   hmiStns[1].wip[14].pnCode[4] := 0;
   hmiStns[1].wip[14].pnCode[5] := 0;
   hmiStns[1].wip[14].pnCode[6] := 0;
   hmiStns[1].wip[14].pnCode[7] := 0;
   hmiStns[1].wip[15].wipCode := -1;
   hmiStns[1].wip[15].pnCode[0] := 0;
   hmiStns[1].wip[15].pnCode[1] := 0;
   hmiStns[1].wip[15].pnCode[2] := 0;
   hmiStns[1].wip[15].pnCode[3] := 0;
   hmiStns[1].wip[15].pnCode[4] := 0;
   hmiStns[1].wip[15].pnCode[5] := 0;
   hmiStns[1].wip[15].pnCode[6] := 0;
   hmiStns[1].wip[15].pnCode[7] := 0;
   hmiStns[1].wip[16].wipCode := -1;
   hmiStns[1].wip[16].pnCode[0] := 0;
   hmiStns[1].wip[16].pnCode[1] := 0;
   hmiStns[1].wip[16].pnCode[2] := 0;
   hmiStns[1].wip[16].pnCode[3] := 0;
   hmiStns[1].wip[16].pnCode[4] := 0;
   hmiStns[1].wip[16].pnCode[5] := 0;
   hmiStns[1].wip[16].pnCode[6] := 0;
   hmiStns[1].wip[16].pnCode[7] := 0;
   hmiStns[1].wip[17].wipCode := -1;
   hmiStns[1].wip[17].pnCode[0] := 0;
   hmiStns[1].wip[17].pnCode[1] := 0;
   hmiStns[1].wip[17].pnCode[2] := 0;
   hmiStns[1].wip[17].pnCode[3] := 0;
   hmiStns[1].wip[17].pnCode[4] := 0;
   hmiStns[1].wip[17].pnCode[5] := 0;
   hmiStns[1].wip[17].pnCode[6] := 0;
   hmiStns[1].wip[17].pnCode[7] := 0;
   hmiStns[1].wip[18].wipCode := -1;
   hmiStns[1].wip[18].pnCode[0] := 0;
   hmiStns[1].wip[18].pnCode[1] := 0;
   hmiStns[1].wip[18].pnCode[2] := 0;
   hmiStns[1].wip[18].pnCode[3] := 0;
   hmiStns[1].wip[18].pnCode[4] := 0;
   hmiStns[1].wip[18].pnCode[5] := 0;
   hmiStns[1].wip[18].pnCode[6] := 0;
   hmiStns[1].wip[18].pnCode[7] := 0;
   hmiStns[1].wip[19].wipCode := -1;
   hmiStns[1].wip[19].pnCode[0] := 0;
   hmiStns[1].wip[19].pnCode[1] := 0;
   hmiStns[1].wip[19].pnCode[2] := 0;
   hmiStns[1].wip[19].pnCode[3] := 0;
   hmiStns[1].wip[19].pnCode[4] := 0;
   hmiStns[1].wip[19].pnCode[5] := 0;
   hmiStns[1].wip[19].pnCode[6] := 0;
   hmiStns[1].wip[19].pnCode[7] := 0;
   hmiStns[1].wip[20].wipCode := -1;
   hmiStns[1].wip[20].pnCode[0] := 0;
   hmiStns[1].wip[20].pnCode[1] := 0;
   hmiStns[1].wip[20].pnCode[2] := 0;
   hmiStns[1].wip[20].pnCode[3] := 0;
   hmiStns[1].wip[20].pnCode[4] := 0;
   hmiStns[1].wip[20].pnCode[5] := 0;
   hmiStns[1].wip[20].pnCode[6] := 0;
   hmiStns[1].wip[20].pnCode[7] := 0;
   hmiStns[1].wip[21].wipCode := -1;
   hmiStns[1].wip[21].pnCode[0] := 0;
   hmiStns[1].wip[21].pnCode[1] := 0;
   hmiStns[1].wip[21].pnCode[2] := 0;
   hmiStns[1].wip[21].pnCode[3] := 0;
   hmiStns[1].wip[21].pnCode[4] := 0;
   hmiStns[1].wip[21].pnCode[5] := 0;
   hmiStns[1].wip[21].pnCode[6] := 0;
   hmiStns[1].wip[21].pnCode[7] := 0;
   hmiStns[1].wip[22].wipCode := -1;
   hmiStns[1].wip[22].pnCode[0] := 0;
   hmiStns[1].wip[22].pnCode[1] := 0;
   hmiStns[1].wip[22].pnCode[2] := 0;
   hmiStns[1].wip[22].pnCode[3] := 0;
   hmiStns[1].wip[22].pnCode[4] := 0;
   hmiStns[1].wip[22].pnCode[5] := 0;
   hmiStns[1].wip[22].pnCode[6] := 0;
   hmiStns[1].wip[22].pnCode[7] := 0;
   hmiStns[1].wip[23].wipCode := -1;
   hmiStns[1].wip[23].pnCode[0] := 0;
   hmiStns[1].wip[23].pnCode[1] := 0;
   hmiStns[1].wip[23].pnCode[2] := 0;
   hmiStns[1].wip[23].pnCode[3] := 0;
   hmiStns[1].wip[23].pnCode[4] := 0;
   hmiStns[1].wip[23].pnCode[5] := 0;
   hmiStns[1].wip[23].pnCode[6] := 0;
   hmiStns[1].wip[23].pnCode[7] := 0;
   hmiStns[1].wip[24].wipCode := -1;
   hmiStns[1].wip[24].pnCode[0] := 0;
   hmiStns[1].wip[24].pnCode[1] := 0;
   hmiStns[1].wip[24].pnCode[2] := 0;
   hmiStns[1].wip[24].pnCode[3] := 0;
   hmiStns[1].wip[24].pnCode[4] := 0;
   hmiStns[1].wip[24].pnCode[5] := 0;
   hmiStns[1].wip[24].pnCode[6] := 0;
   hmiStns[1].wip[24].pnCode[7] := 0;
   hmiStns[1].wip[25].wipCode := -1;
   hmiStns[1].wip[25].pnCode[0] := 0;
   hmiStns[1].wip[25].pnCode[1] := 0;
   hmiStns[1].wip[25].pnCode[2] := 0;
   hmiStns[1].wip[25].pnCode[3] := 0;
   hmiStns[1].wip[25].pnCode[4] := 0;
   hmiStns[1].wip[25].pnCode[5] := 0;
   hmiStns[1].wip[25].pnCode[6] := 0;
   hmiStns[1].wip[25].pnCode[7] := 0;
   hmiStns[1].wip[26].wipCode := -1;
   hmiStns[1].wip[26].pnCode[0] := 0;
   hmiStns[1].wip[26].pnCode[1] := 0;
   hmiStns[1].wip[26].pnCode[2] := 0;
   hmiStns[1].wip[26].pnCode[3] := 0;
   hmiStns[1].wip[26].pnCode[4] := 0;
   hmiStns[1].wip[26].pnCode[5] := 0;
   hmiStns[1].wip[26].pnCode[6] := 0;
   hmiStns[1].wip[26].pnCode[7] := 0;
   hmiStns[1].wip[27].wipCode := -1;
   hmiStns[1].wip[27].pnCode[0] := 0;
   hmiStns[1].wip[27].pnCode[1] := 0;
   hmiStns[1].wip[27].pnCode[2] := 0;
   hmiStns[1].wip[27].pnCode[3] := 0;
   hmiStns[1].wip[27].pnCode[4] := 0;
   hmiStns[1].wip[27].pnCode[5] := 0;
   hmiStns[1].wip[27].pnCode[6] := 0;
   hmiStns[1].wip[27].pnCode[7] := 0;
   hmiStns[1].wip[28].wipCode := -1;
   hmiStns[1].wip[28].pnCode[0] := 0;
   hmiStns[1].wip[28].pnCode[1] := 0;
   hmiStns[1].wip[28].pnCode[2] := 0;
   hmiStns[1].wip[28].pnCode[3] := 0;
   hmiStns[1].wip[28].pnCode[4] := 0;
   hmiStns[1].wip[28].pnCode[5] := 0;
   hmiStns[1].wip[28].pnCode[6] := 0;
   hmiStns[1].wip[28].pnCode[7] := 0;
   hmiStns[1].wip[29].wipCode := -1;
   hmiStns[1].wip[29].pnCode[0] := 0;
   hmiStns[1].wip[29].pnCode[1] := 0;
   hmiStns[1].wip[29].pnCode[2] := 0;
   hmiStns[1].wip[29].pnCode[3] := 0;
   hmiStns[1].wip[29].pnCode[4] := 0;
   hmiStns[1].wip[29].pnCode[5] := 0;
   hmiStns[1].wip[29].pnCode[6] := 0;
   hmiStns[1].wip[29].pnCode[7] := 0;
   hmiStns[1].wip[30].wipCode := -1;
   hmiStns[1].wip[30].pnCode[0] := 0;
   hmiStns[1].wip[30].pnCode[1] := 0;
   hmiStns[1].wip[30].pnCode[2] := 0;
   hmiStns[1].wip[30].pnCode[3] := 0;
   hmiStns[1].wip[30].pnCode[4] := 0;
   hmiStns[1].wip[30].pnCode[5] := 0;
   hmiStns[1].wip[30].pnCode[6] := 0;
   hmiStns[1].wip[30].pnCode[7] := 0;
   hmiStns[1].wip[31].wipCode := -1;
   hmiStns[1].wip[31].pnCode[0] := 0;
   hmiStns[1].wip[31].pnCode[1] := 0;
   hmiStns[1].wip[31].pnCode[2] := 0;
   hmiStns[1].wip[31].pnCode[3] := 0;
   hmiStns[1].wip[31].pnCode[4] := 0;
   hmiStns[1].wip[31].pnCode[5] := 0;
   hmiStns[1].wip[31].pnCode[6] := 0;
   hmiStns[1].wip[31].pnCode[7] := 0;
   hmiStns[1].wip[32].wipCode := -1;
   hmiStns[1].wip[32].pnCode[0] := 0;
   hmiStns[1].wip[32].pnCode[1] := 0;
   hmiStns[1].wip[32].pnCode[2] := 0;
   hmiStns[1].wip[32].pnCode[3] := 0;
   hmiStns[1].wip[32].pnCode[4] := 0;
   hmiStns[1].wip[32].pnCode[5] := 0;
   hmiStns[1].wip[32].pnCode[6] := 0;
   hmiStns[1].wip[32].pnCode[7] := 0;
   hmiStns[1].wip[33].wipCode := -1;
   hmiStns[1].wip[33].pnCode[0] := 0;
   hmiStns[1].wip[33].pnCode[1] := 0;
   hmiStns[1].wip[33].pnCode[2] := 0;
   hmiStns[1].wip[33].pnCode[3] := 0;
   hmiStns[1].wip[33].pnCode[4] := 0;
   hmiStns[1].wip[33].pnCode[5] := 0;
   hmiStns[1].wip[33].pnCode[6] := 0;
   hmiStns[1].wip[33].pnCode[7] := 0;
   hmiStns[1].wip[34].wipCode := -1;
   hmiStns[1].wip[34].pnCode[0] := 0;
   hmiStns[1].wip[34].pnCode[1] := 0;
   hmiStns[1].wip[34].pnCode[2] := 0;
   hmiStns[1].wip[34].pnCode[3] := 0;
   hmiStns[1].wip[34].pnCode[4] := 0;
   hmiStns[1].wip[34].pnCode[5] := 0;
   hmiStns[1].wip[34].pnCode[6] := 0;
   hmiStns[1].wip[34].pnCode[7] := 0;
   hmiStns[1].wip[35].wipCode := -1;
   hmiStns[1].wip[35].pnCode[0] := 0;
   hmiStns[1].wip[35].pnCode[1] := 0;
   hmiStns[1].wip[35].pnCode[2] := 0;
   hmiStns[1].wip[35].pnCode[3] := 0;
   hmiStns[1].wip[35].pnCode[4] := 0;
   hmiStns[1].wip[35].pnCode[5] := 0;
   hmiStns[1].wip[35].pnCode[6] := 0;
   hmiStns[1].wip[35].pnCode[7] := 0;
   hmiStns[1].wip[36].wipCode := -1;
   hmiStns[1].wip[36].pnCode[0] := 0;
   hmiStns[1].wip[36].pnCode[1] := 0;
   hmiStns[1].wip[36].pnCode[2] := 0;
   hmiStns[1].wip[36].pnCode[3] := 0;
   hmiStns[1].wip[36].pnCode[4] := 0;
   hmiStns[1].wip[36].pnCode[5] := 0;
   hmiStns[1].wip[36].pnCode[6] := 0;
   hmiStns[1].wip[36].pnCode[7] := 0;
   hmiStns[1].wip[37].wipCode := -1;
   hmiStns[1].wip[37].pnCode[0] := 0;
   hmiStns[1].wip[37].pnCode[1] := 0;
   hmiStns[1].wip[37].pnCode[2] := 0;
   hmiStns[1].wip[37].pnCode[3] := 0;
   hmiStns[1].wip[37].pnCode[4] := 0;
   hmiStns[1].wip[37].pnCode[5] := 0;
   hmiStns[1].wip[37].pnCode[6] := 0;
   hmiStns[1].wip[37].pnCode[7] := 0;
   hmiStns[1].wip[38].wipCode := -1;
   hmiStns[1].wip[38].pnCode[0] := 0;
   hmiStns[1].wip[38].pnCode[1] := 0;
   hmiStns[1].wip[38].pnCode[2] := 0;
   hmiStns[1].wip[38].pnCode[3] := 0;
   hmiStns[1].wip[38].pnCode[4] := 0;
   hmiStns[1].wip[38].pnCode[5] := 0;
   hmiStns[1].wip[38].pnCode[6] := 0;
   hmiStns[1].wip[38].pnCode[7] := 0;
   hmiStns[1].wip[39].wipCode := -1;
   hmiStns[1].wip[39].pnCode[0] := 0;
   hmiStns[1].wip[39].pnCode[1] := 0;
   hmiStns[1].wip[39].pnCode[2] := 0;
   hmiStns[1].wip[39].pnCode[3] := 0;
   hmiStns[1].wip[39].pnCode[4] := 0;
   hmiStns[1].wip[39].pnCode[5] := 0;
   hmiStns[1].wip[39].pnCode[6] := 0;
   hmiStns[1].wip[39].pnCode[7] := 0;
   hmiStns[1].wip[40].wipCode := -1;
   hmiStns[1].wip[40].pnCode[0] := 0;
   hmiStns[1].wip[40].pnCode[1] := 0;
   hmiStns[1].wip[40].pnCode[2] := 0;
   hmiStns[1].wip[40].pnCode[3] := 0;
   hmiStns[1].wip[40].pnCode[4] := 0;
   hmiStns[1].wip[40].pnCode[5] := 0;
   hmiStns[1].wip[40].pnCode[6] := 0;
   hmiStns[1].wip[40].pnCode[7] := 0;
   hmiStns[1].wip[41].wipCode := -1;
   hmiStns[1].wip[41].pnCode[0] := 0;
   hmiStns[1].wip[41].pnCode[1] := 0;
   hmiStns[1].wip[41].pnCode[2] := 0;
   hmiStns[1].wip[41].pnCode[3] := 0;
   hmiStns[1].wip[41].pnCode[4] := 0;
   hmiStns[1].wip[41].pnCode[5] := 0;
   hmiStns[1].wip[41].pnCode[6] := 0;
   hmiStns[1].wip[41].pnCode[7] := 0;
   hmiStns[1].wip[42].wipCode := -1;
   hmiStns[1].wip[42].pnCode[0] := 0;
   hmiStns[1].wip[42].pnCode[1] := 0;
   hmiStns[1].wip[42].pnCode[2] := 0;
   hmiStns[1].wip[42].pnCode[3] := 0;
   hmiStns[1].wip[42].pnCode[4] := 0;
   hmiStns[1].wip[42].pnCode[5] := 0;
   hmiStns[1].wip[42].pnCode[6] := 0;
   hmiStns[1].wip[42].pnCode[7] := 0;
   hmiStns[1].wip[43].wipCode := -1;
   hmiStns[1].wip[43].pnCode[0] := 0;
   hmiStns[1].wip[43].pnCode[1] := 0;
   hmiStns[1].wip[43].pnCode[2] := 0;
   hmiStns[1].wip[43].pnCode[3] := 0;
   hmiStns[1].wip[43].pnCode[4] := 0;
   hmiStns[1].wip[43].pnCode[5] := 0;
   hmiStns[1].wip[43].pnCode[6] := 0;
   hmiStns[1].wip[43].pnCode[7] := 0;
   hmiStns[1].wip[44].wipCode := -1;
   hmiStns[1].wip[44].pnCode[0] := 0;
   hmiStns[1].wip[44].pnCode[1] := 0;
   hmiStns[1].wip[44].pnCode[2] := 0;
   hmiStns[1].wip[44].pnCode[3] := 0;
   hmiStns[1].wip[44].pnCode[4] := 0;
   hmiStns[1].wip[44].pnCode[5] := 0;
   hmiStns[1].wip[44].pnCode[6] := 0;
   hmiStns[1].wip[44].pnCode[7] := 0;
   hmiStns[1].wip[45].wipCode := -1;
   hmiStns[1].wip[45].pnCode[0] := 0;
   hmiStns[1].wip[45].pnCode[1] := 0;
   hmiStns[1].wip[45].pnCode[2] := 0;
   hmiStns[1].wip[45].pnCode[3] := 0;
   hmiStns[1].wip[45].pnCode[4] := 0;
   hmiStns[1].wip[45].pnCode[5] := 0;
   hmiStns[1].wip[45].pnCode[6] := 0;
   hmiStns[1].wip[45].pnCode[7] := 0;
   hmiStns[1].wip[46].wipCode := -1;
   hmiStns[1].wip[46].pnCode[0] := 0;
   hmiStns[1].wip[46].pnCode[1] := 0;
   hmiStns[1].wip[46].pnCode[2] := 0;
   hmiStns[1].wip[46].pnCode[3] := 0;
   hmiStns[1].wip[46].pnCode[4] := 0;
   hmiStns[1].wip[46].pnCode[5] := 0;
   hmiStns[1].wip[46].pnCode[6] := 0;
   hmiStns[1].wip[46].pnCode[7] := 0;
   hmiStns[1].wip[47].wipCode := -1;
   hmiStns[1].wip[47].pnCode[0] := 0;
   hmiStns[1].wip[47].pnCode[1] := 0;
   hmiStns[1].wip[47].pnCode[2] := 0;
   hmiStns[1].wip[47].pnCode[3] := 0;
   hmiStns[1].wip[47].pnCode[4] := 0;
   hmiStns[1].wip[47].pnCode[5] := 0;
   hmiStns[1].wip[47].pnCode[6] := 0;
   hmiStns[1].wip[47].pnCode[7] := 0;
   hmiStns[1].wip[48].wipCode := -1;
   hmiStns[1].wip[48].pnCode[0] := 0;
   hmiStns[1].wip[48].pnCode[1] := 0;
   hmiStns[1].wip[48].pnCode[2] := 0;
   hmiStns[1].wip[48].pnCode[3] := 0;
   hmiStns[1].wip[48].pnCode[4] := 0;
   hmiStns[1].wip[48].pnCode[5] := 0;
   hmiStns[1].wip[48].pnCode[6] := 0;
   hmiStns[1].wip[48].pnCode[7] := 0;
   hmiStns[1].wip[49].wipCode := -1;
   hmiStns[1].wip[49].pnCode[0] := 0;
   hmiStns[1].wip[49].pnCode[1] := 0;
   hmiStns[1].wip[49].pnCode[2] := 0;
   hmiStns[1].wip[49].pnCode[3] := 0;
   hmiStns[1].wip[49].pnCode[4] := 0;
   hmiStns[1].wip[49].pnCode[5] := 0;
   hmiStns[1].wip[49].pnCode[6] := 0;
   hmiStns[1].wip[49].pnCode[7] := 0;
   hmiStns[2].wip[0].wipCode := 53014;
   hmiStns[2].wip[0].pnCode[0] := 0;
   hmiStns[2].wip[0].pnCode[1] := 243000;
   hmiStns[2].wip[0].pnCode[2] := 148000;
   hmiStns[2].wip[0].pnCode[3] := 0;
   hmiStns[2].wip[0].pnCode[4] := 0;
   hmiStns[2].wip[0].pnCode[5] := 0;
   hmiStns[2].wip[0].pnCode[6] := 147000;
   hmiStns[2].wip[0].pnCode[7] := 149000;
   hmiStns[2].wip[1].wipCode := 19031;
   hmiStns[2].wip[1].pnCode[0] := 0;
   hmiStns[2].wip[1].pnCode[1] := 243000;
   hmiStns[2].wip[1].pnCode[2] := 53000;
   hmiStns[2].wip[1].pnCode[3] := 0;
   hmiStns[2].wip[1].pnCode[4] := 0;
   hmiStns[2].wip[1].pnCode[5] := 0;
   hmiStns[2].wip[1].pnCode[6] := 31000;
   hmiStns[2].wip[1].pnCode[7] := 71000;
   hmiStns[2].wip[2].wipCode := 21028;
   hmiStns[2].wip[2].pnCode[0] := 0;
   hmiStns[2].wip[2].pnCode[1] := 243000;
   hmiStns[2].wip[2].pnCode[2] := 57000;
   hmiStns[2].wip[2].pnCode[3] := 0;
   hmiStns[2].wip[2].pnCode[4] := 0;
   hmiStns[2].wip[2].pnCode[5] := 0;
   hmiStns[2].wip[2].pnCode[6] := 25000;
   hmiStns[2].wip[2].pnCode[7] := 18000;
   hmiStns[2].wip[3].wipCode := 22008;
   hmiStns[2].wip[3].pnCode[0] := 0;
   hmiStns[2].wip[3].pnCode[1] := 243000;
   hmiStns[2].wip[3].pnCode[2] := 84000;
   hmiStns[2].wip[3].pnCode[3] := 0;
   hmiStns[2].wip[3].pnCode[4] := 0;
   hmiStns[2].wip[3].pnCode[5] := 0;
   hmiStns[2].wip[3].pnCode[6] := 31000;
   hmiStns[2].wip[3].pnCode[7] := 71000;
   hmiStns[2].wip[4].wipCode := 20050;
   hmiStns[2].wip[4].pnCode[0] := 0;
   hmiStns[2].wip[4].pnCode[1] := 243000;
   hmiStns[2].wip[4].pnCode[2] := 70000;
   hmiStns[2].wip[4].pnCode[3] := 72000;
   hmiStns[2].wip[4].pnCode[4] := 0;
   hmiStns[2].wip[4].pnCode[5] := 58000;
   hmiStns[2].wip[4].pnCode[6] := 33000;
   hmiStns[2].wip[4].pnCode[7] := 73000;
   hmiStns[2].wip[5].wipCode := 27040;
   hmiStns[2].wip[5].pnCode[0] := 0;
   hmiStns[2].wip[5].pnCode[1] := 243000;
   hmiStns[2].wip[5].pnCode[2] := 127000;
   hmiStns[2].wip[5].pnCode[3] := 0;
   hmiStns[2].wip[5].pnCode[4] := 0;
   hmiStns[2].wip[5].pnCode[5] := 100000;
   hmiStns[2].wip[5].pnCode[6] := 101000;
   hmiStns[2].wip[5].pnCode[7] := 128000;
   hmiStns[2].wip[6].wipCode := 28041;
   hmiStns[2].wip[6].pnCode[0] := 0;
   hmiStns[2].wip[6].pnCode[1] := 243000;
   hmiStns[2].wip[6].pnCode[2] := 122000;
   hmiStns[2].wip[6].pnCode[3] := 123000;
   hmiStns[2].wip[6].pnCode[4] := 0;
   hmiStns[2].wip[6].pnCode[5] := 102000;
   hmiStns[2].wip[6].pnCode[6] := 103000;
   hmiStns[2].wip[6].pnCode[7] := 133000;
   hmiStns[2].wip[7].wipCode := 29044;
   hmiStns[2].wip[7].pnCode[0] := 0;
   hmiStns[2].wip[7].pnCode[1] := 243000;
   hmiStns[2].wip[7].pnCode[2] := 100000;
   hmiStns[2].wip[7].pnCode[3] := 128000;
   hmiStns[2].wip[7].pnCode[4] := 0;
   hmiStns[2].wip[7].pnCode[5] := 102000;
   hmiStns[2].wip[7].pnCode[6] := 104000;
   hmiStns[2].wip[7].pnCode[7] := 133000;
   hmiStns[2].wip[8].wipCode := 30041;
   hmiStns[2].wip[8].pnCode[0] := 0;
   hmiStns[2].wip[8].pnCode[1] := 243000;
   hmiStns[2].wip[8].pnCode[2] := 105000;
   hmiStns[2].wip[8].pnCode[3] := 123000;
   hmiStns[2].wip[8].pnCode[4] := 0;
   hmiStns[2].wip[8].pnCode[5] := 106000;
   hmiStns[2].wip[8].pnCode[6] := 107000;
   hmiStns[2].wip[8].pnCode[7] := 133000;
   hmiStns[2].wip[9].wipCode := 31040;
   hmiStns[2].wip[9].pnCode[0] := 0;
   hmiStns[2].wip[9].pnCode[1] := 243000;
   hmiStns[2].wip[9].pnCode[2] := 100000;
   hmiStns[2].wip[9].pnCode[3] := 0;
   hmiStns[2].wip[9].pnCode[4] := 0;
   hmiStns[2].wip[9].pnCode[5] := 127000;
   hmiStns[2].wip[9].pnCode[6] := 107000;
   hmiStns[2].wip[9].pnCode[7] := 128000;
   hmiStns[2].wip[10].wipCode := 32043;
   hmiStns[2].wip[10].pnCode[0] := 0;
   hmiStns[2].wip[10].pnCode[1] := 243000;
   hmiStns[2].wip[10].pnCode[2] := 100000;
   hmiStns[2].wip[10].pnCode[3] := 128000;
   hmiStns[2].wip[10].pnCode[4] := 0;
   hmiStns[2].wip[10].pnCode[5] := 106000;
   hmiStns[2].wip[10].pnCode[6] := 107000;
   hmiStns[2].wip[10].pnCode[7] := 123000;
   hmiStns[2].wip[11].wipCode := 33043;
   hmiStns[2].wip[11].pnCode[0] := 0;
   hmiStns[2].wip[11].pnCode[1] := 243000;
   hmiStns[2].wip[11].pnCode[2] := 108000;
   hmiStns[2].wip[11].pnCode[3] := 0;
   hmiStns[2].wip[11].pnCode[4] := 0;
   hmiStns[2].wip[11].pnCode[5] := 0;
   hmiStns[2].wip[11].pnCode[6] := 107000;
   hmiStns[2].wip[11].pnCode[7] := 109000;
   hmiStns[2].wip[12].wipCode := 34036;
   hmiStns[2].wip[12].pnCode[0] := 0;
   hmiStns[2].wip[12].pnCode[1] := 243000;
   hmiStns[2].wip[12].pnCode[2] := 110000;
   hmiStns[2].wip[12].pnCode[3] := 113000;
   hmiStns[2].wip[12].pnCode[4] := 0;
   hmiStns[2].wip[12].pnCode[5] := 112000;
   hmiStns[2].wip[12].pnCode[6] := 114000;
   hmiStns[2].wip[12].pnCode[7] := 111000;
   hmiStns[2].wip[13].wipCode := 35037;
   hmiStns[2].wip[13].pnCode[0] := 0;
   hmiStns[2].wip[13].pnCode[1] := 243000;
   hmiStns[2].wip[13].pnCode[2] := 115000;
   hmiStns[2].wip[13].pnCode[3] := 0;
   hmiStns[2].wip[13].pnCode[4] := 0;
   hmiStns[2].wip[13].pnCode[5] := 112000;
   hmiStns[2].wip[13].pnCode[6] := 114000;
   hmiStns[2].wip[13].pnCode[7] := 113000;
   hmiStns[2].wip[14].wipCode := 36038;
   hmiStns[2].wip[14].pnCode[0] := 0;
   hmiStns[2].wip[14].pnCode[1] := 243000;
   hmiStns[2].wip[14].pnCode[2] := 116000;
   hmiStns[2].wip[14].pnCode[3] := 111000;
   hmiStns[2].wip[14].pnCode[4] := 0;
   hmiStns[2].wip[14].pnCode[5] := 118000;
   hmiStns[2].wip[14].pnCode[6] := 114000;
   hmiStns[2].wip[14].pnCode[7] := 117000;
   hmiStns[2].wip[15].wipCode := 37038;
   hmiStns[2].wip[15].pnCode[0] := 0;
   hmiStns[2].wip[15].pnCode[1] := 243000;
   hmiStns[2].wip[15].pnCode[2] := 116000;
   hmiStns[2].wip[15].pnCode[3] := 117000;
   hmiStns[2].wip[15].pnCode[4] := 0;
   hmiStns[2].wip[15].pnCode[5] := 118000;
   hmiStns[2].wip[15].pnCode[6] := 120000;
   hmiStns[2].wip[15].pnCode[7] := 111000;
   hmiStns[2].wip[16].wipCode := 38039;
   hmiStns[2].wip[16].pnCode[0] := 0;
   hmiStns[2].wip[16].pnCode[1] := 243000;
   hmiStns[2].wip[16].pnCode[2] := 119000;
   hmiStns[2].wip[16].pnCode[3] := 0;
   hmiStns[2].wip[16].pnCode[4] := 0;
   hmiStns[2].wip[16].pnCode[5] := 121000;
   hmiStns[2].wip[16].pnCode[6] := 114000;
   hmiStns[2].wip[16].pnCode[7] := 111000;
   hmiStns[2].wip[17].wipCode := 39042;
   hmiStns[2].wip[17].pnCode[0] := 0;
   hmiStns[2].wip[17].pnCode[1] := 243000;
   hmiStns[2].wip[17].pnCode[2] := 124000;
   hmiStns[2].wip[17].pnCode[3] := 125000;
   hmiStns[2].wip[17].pnCode[4] := 0;
   hmiStns[2].wip[17].pnCode[5] := 122000;
   hmiStns[2].wip[17].pnCode[6] := 107000;
   hmiStns[2].wip[17].pnCode[7] := 123000;
   hmiStns[2].wip[18].wipCode := 40040;
   hmiStns[2].wip[18].pnCode[0] := 0;
   hmiStns[2].wip[18].pnCode[1] := 243000;
   hmiStns[2].wip[18].pnCode[2] := 100000;
   hmiStns[2].wip[18].pnCode[3] := 0;
   hmiStns[2].wip[18].pnCode[4] := 0;
   hmiStns[2].wip[18].pnCode[5] := 127000;
   hmiStns[2].wip[18].pnCode[6] := 126000;
   hmiStns[2].wip[18].pnCode[7] := 128000;
   hmiStns[2].wip[19].wipCode := 41045;
   hmiStns[2].wip[19].pnCode[0] := 0;
   hmiStns[2].wip[19].pnCode[1] := 243000;
   hmiStns[2].wip[19].pnCode[2] := 127000;
   hmiStns[2].wip[19].pnCode[3] := 123000;
   hmiStns[2].wip[19].pnCode[4] := 0;
   hmiStns[2].wip[19].pnCode[5] := 122000;
   hmiStns[2].wip[19].pnCode[6] := 129000;
   hmiStns[2].wip[19].pnCode[7] := 128000;
   hmiStns[2].wip[20].wipCode := 42044;
   hmiStns[2].wip[20].pnCode[0] := 0;
   hmiStns[2].wip[20].pnCode[1] := 243000;
   hmiStns[2].wip[20].pnCode[2] := 130000;
   hmiStns[2].wip[20].pnCode[3] := 0;
   hmiStns[2].wip[20].pnCode[4] := 0;
   hmiStns[2].wip[20].pnCode[5] := 0;
   hmiStns[2].wip[20].pnCode[6] := 126000;
   hmiStns[2].wip[20].pnCode[7] := 131000;
   hmiStns[2].wip[21].wipCode := 44019;
   hmiStns[2].wip[21].pnCode[0] := 0;
   hmiStns[2].wip[21].pnCode[1] := 243000;
   hmiStns[2].wip[21].pnCode[2] := 132000;
   hmiStns[2].wip[21].pnCode[3] := 0;
   hmiStns[2].wip[21].pnCode[4] := 0;
   hmiStns[2].wip[21].pnCode[5] := 0;
   hmiStns[2].wip[21].pnCode[6] := 143000;
   hmiStns[2].wip[21].pnCode[7] := 133000;
   hmiStns[2].wip[22].wipCode := 45017;
   hmiStns[2].wip[22].pnCode[0] := 0;
   hmiStns[2].wip[22].pnCode[1] := 243000;
   hmiStns[2].wip[22].pnCode[2] := 134000;
   hmiStns[2].wip[22].pnCode[3] := 0;
   hmiStns[2].wip[22].pnCode[4] := 0;
   hmiStns[2].wip[22].pnCode[5] := 0;
   hmiStns[2].wip[22].pnCode[6] := 143000;
   hmiStns[2].wip[22].pnCode[7] := 135000;
   hmiStns[2].wip[23].wipCode := 46018;
   hmiStns[2].wip[23].pnCode[0] := 0;
   hmiStns[2].wip[23].pnCode[1] := 243000;
   hmiStns[2].wip[23].pnCode[2] := 142000;
   hmiStns[2].wip[23].pnCode[3] := 0;
   hmiStns[2].wip[23].pnCode[4] := 0;
   hmiStns[2].wip[23].pnCode[5] := 0;
   hmiStns[2].wip[23].pnCode[6] := 143000;
   hmiStns[2].wip[23].pnCode[7] := 133000;
   hmiStns[2].wip[24].wipCode := 47017;
   hmiStns[2].wip[24].pnCode[0] := 0;
   hmiStns[2].wip[24].pnCode[1] := 243000;
   hmiStns[2].wip[24].pnCode[2] := 136000;
   hmiStns[2].wip[24].pnCode[3] := 0;
   hmiStns[2].wip[24].pnCode[4] := 0;
   hmiStns[2].wip[24].pnCode[5] := 0;
   hmiStns[2].wip[24].pnCode[6] := 143000;
   hmiStns[2].wip[24].pnCode[7] := 135000;
   hmiStns[2].wip[25].wipCode := 48021;
   hmiStns[2].wip[25].pnCode[0] := 0;
   hmiStns[2].wip[25].pnCode[1] := 243000;
   hmiStns[2].wip[25].pnCode[2] := 137000;
   hmiStns[2].wip[25].pnCode[3] := 0;
   hmiStns[2].wip[25].pnCode[4] := 0;
   hmiStns[2].wip[25].pnCode[5] := 0;
   hmiStns[2].wip[25].pnCode[6] := 140000;
   hmiStns[2].wip[25].pnCode[7] := 128000;
   hmiStns[2].wip[26].wipCode := 49022;
   hmiStns[2].wip[26].pnCode[0] := 0;
   hmiStns[2].wip[26].pnCode[1] := 243000;
   hmiStns[2].wip[26].pnCode[2] := 138000;
   hmiStns[2].wip[26].pnCode[3] := 0;
   hmiStns[2].wip[26].pnCode[4] := 0;
   hmiStns[2].wip[26].pnCode[5] := 0;
   hmiStns[2].wip[26].pnCode[6] := 140000;
   hmiStns[2].wip[26].pnCode[7] := 139000;
   hmiStns[2].wip[27].wipCode := 50020;
   hmiStns[2].wip[27].pnCode[0] := 0;
   hmiStns[2].wip[27].pnCode[1] := 243000;
   hmiStns[2].wip[27].pnCode[2] := 141000;
   hmiStns[2].wip[27].pnCode[3] := 0;
   hmiStns[2].wip[27].pnCode[4] := 0;
   hmiStns[2].wip[27].pnCode[5] := 0;
   hmiStns[2].wip[27].pnCode[6] := 140000;
   hmiStns[2].wip[27].pnCode[7] := 125000;
   hmiStns[2].wip[28].wipCode := 51013;
   hmiStns[2].wip[28].pnCode[0] := 0;
   hmiStns[2].wip[28].pnCode[1] := 243000;
   hmiStns[2].wip[28].pnCode[2] := 148000;
   hmiStns[2].wip[28].pnCode[3] := 0;
   hmiStns[2].wip[28].pnCode[4] := 0;
   hmiStns[2].wip[28].pnCode[5] := 0;
   hmiStns[2].wip[28].pnCode[6] := 144000;
   hmiStns[2].wip[28].pnCode[7] := 149000;
   hmiStns[2].wip[29].wipCode := 52016;
   hmiStns[2].wip[29].pnCode[0] := 0;
   hmiStns[2].wip[29].pnCode[1] := 243000;
   hmiStns[2].wip[29].pnCode[2] := 145000;
   hmiStns[2].wip[29].pnCode[3] := 0;
   hmiStns[2].wip[29].pnCode[4] := 0;
   hmiStns[2].wip[29].pnCode[5] := 0;
   hmiStns[2].wip[29].pnCode[6] := 147000;
   hmiStns[2].wip[29].pnCode[7] := 146000;
   hmiStns[2].wip[30].wipCode := 54012;
   hmiStns[2].wip[30].pnCode[0] := 0;
   hmiStns[2].wip[30].pnCode[1] := 243000;
   hmiStns[2].wip[30].pnCode[2] := 159000;
   hmiStns[2].wip[30].pnCode[3] := 0;
   hmiStns[2].wip[30].pnCode[4] := 0;
   hmiStns[2].wip[30].pnCode[5] := 0;
   hmiStns[2].wip[30].pnCode[6] := 144000;
   hmiStns[2].wip[30].pnCode[7] := 160000;
   hmiStns[2].wip[31].wipCode := 55014;
   hmiStns[2].wip[31].pnCode[0] := 0;
   hmiStns[2].wip[31].pnCode[1] := 243000;
   hmiStns[2].wip[31].pnCode[2] := 163000;
   hmiStns[2].wip[31].pnCode[3] := 0;
   hmiStns[2].wip[31].pnCode[4] := 0;
   hmiStns[2].wip[31].pnCode[5] := 0;
   hmiStns[2].wip[31].pnCode[6] := 147000;
   hmiStns[2].wip[31].pnCode[7] := 146000;
   hmiStns[2].wip[32].wipCode := 56012;
   hmiStns[2].wip[32].pnCode[0] := 0;
   hmiStns[2].wip[32].pnCode[1] := 243000;
   hmiStns[2].wip[32].pnCode[2] := 159000;
   hmiStns[2].wip[32].pnCode[3] := 0;
   hmiStns[2].wip[32].pnCode[4] := 0;
   hmiStns[2].wip[32].pnCode[5] := 0;
   hmiStns[2].wip[32].pnCode[6] := 147000;
   hmiStns[2].wip[32].pnCode[7] := 160000;
   hmiStns[2].wip[33].wipCode := 57033;
   hmiStns[2].wip[33].pnCode[0] := 0;
   hmiStns[2].wip[33].pnCode[1] := 243000;
   hmiStns[2].wip[33].pnCode[2] := 152000;
   hmiStns[2].wip[33].pnCode[3] := 151000;
   hmiStns[2].wip[33].pnCode[4] := 0;
   hmiStns[2].wip[33].pnCode[5] := 150000;
   hmiStns[2].wip[33].pnCode[6] := 154000;
   hmiStns[2].wip[33].pnCode[7] := 153000;
   hmiStns[2].wip[34].wipCode := 58034;
   hmiStns[2].wip[34].pnCode[0] := 0;
   hmiStns[2].wip[34].pnCode[1] := 243000;
   hmiStns[2].wip[34].pnCode[2] := 152000;
   hmiStns[2].wip[34].pnCode[3] := 0;
   hmiStns[2].wip[34].pnCode[4] := 0;
   hmiStns[2].wip[34].pnCode[5] := 155000;
   hmiStns[2].wip[34].pnCode[6] := 154000;
   hmiStns[2].wip[34].pnCode[7] := 153000;
   hmiStns[2].wip[35].wipCode := 59035;
   hmiStns[2].wip[35].pnCode[0] := 0;
   hmiStns[2].wip[35].pnCode[1] := 243000;
   hmiStns[2].wip[35].pnCode[2] := 156000;
   hmiStns[2].wip[35].pnCode[3] := 0;
   hmiStns[2].wip[35].pnCode[4] := 0;
   hmiStns[2].wip[35].pnCode[5] := 0;
   hmiStns[2].wip[35].pnCode[6] := 154000;
   hmiStns[2].wip[35].pnCode[7] := 157000;
   hmiStns[2].wip[36].wipCode := 60015;
   hmiStns[2].wip[36].pnCode[0] := 0;
   hmiStns[2].wip[36].pnCode[1] := 243000;
   hmiStns[2].wip[36].pnCode[2] := 159000;
   hmiStns[2].wip[36].pnCode[3] := 0;
   hmiStns[2].wip[36].pnCode[4] := 0;
   hmiStns[2].wip[36].pnCode[5] := 0;
   hmiStns[2].wip[36].pnCode[6] := 161000;
   hmiStns[2].wip[36].pnCode[7] := 160000;
   hmiStns[2].wip[37].wipCode := 61014;
   hmiStns[2].wip[37].pnCode[0] := 0;
   hmiStns[2].wip[37].pnCode[1] := 243000;
   hmiStns[2].wip[37].pnCode[2] := 158000;
   hmiStns[2].wip[37].pnCode[3] := 0;
   hmiStns[2].wip[37].pnCode[4] := 0;
   hmiStns[2].wip[37].pnCode[5] := 0;
   hmiStns[2].wip[37].pnCode[6] := 161000;
   hmiStns[2].wip[37].pnCode[7] := 160000;
   hmiStns[2].wip[38].wipCode := 62015;
   hmiStns[2].wip[38].pnCode[0] := 0;
   hmiStns[2].wip[38].pnCode[1] := 243000;
   hmiStns[2].wip[38].pnCode[2] := 162000;
   hmiStns[2].wip[38].pnCode[3] := 0;
   hmiStns[2].wip[38].pnCode[4] := 0;
   hmiStns[2].wip[38].pnCode[5] := 0;
   hmiStns[2].wip[38].pnCode[6] := 161000;
   hmiStns[2].wip[38].pnCode[7] := 160000;
   hmiStns[2].wip[39].wipCode := 63014;
   hmiStns[2].wip[39].pnCode[0] := 0;
   hmiStns[2].wip[39].pnCode[1] := 243000;
   hmiStns[2].wip[39].pnCode[2] := 163000;
   hmiStns[2].wip[39].pnCode[3] := 0;
   hmiStns[2].wip[39].pnCode[4] := 0;
   hmiStns[2].wip[39].pnCode[5] := 0;
   hmiStns[2].wip[39].pnCode[6] := 161000;
   hmiStns[2].wip[39].pnCode[7] := 146000;
   hmiStns[2].wip[40].wipCode := 43051;
   hmiStns[2].wip[40].pnCode[0] := 0;
   hmiStns[2].wip[40].pnCode[1] := 243000;
   hmiStns[2].wip[40].pnCode[2] := 105000;
   hmiStns[2].wip[40].pnCode[3] := 128000;
   hmiStns[2].wip[40].pnCode[4] := 0;
   hmiStns[2].wip[40].pnCode[5] := 127000;
   hmiStns[2].wip[40].pnCode[6] := 126000;
   hmiStns[2].wip[40].pnCode[7] := 133000;
   hmiStns[2].wip[41].wipCode := 75057;
   hmiStns[2].wip[41].pnCode[0] := 0;
   hmiStns[2].wip[41].pnCode[1] := 0;
   hmiStns[2].wip[41].pnCode[2] := 0;
   hmiStns[2].wip[41].pnCode[3] := 0;
   hmiStns[2].wip[41].pnCode[4] := 0;
   hmiStns[2].wip[41].pnCode[5] := 0;
   hmiStns[2].wip[41].pnCode[6] := 0;
   hmiStns[2].wip[41].pnCode[7] := 0;
   hmiStns[2].wip[42].wipCode := -1;
   hmiStns[2].wip[42].pnCode[0] := 0;
   hmiStns[2].wip[42].pnCode[1] := 0;
   hmiStns[2].wip[42].pnCode[2] := 0;
   hmiStns[2].wip[42].pnCode[3] := 0;
   hmiStns[2].wip[42].pnCode[4] := 0;
   hmiStns[2].wip[42].pnCode[5] := 0;
   hmiStns[2].wip[42].pnCode[6] := 0;
   hmiStns[2].wip[42].pnCode[7] := 0;
   hmiStns[2].wip[43].wipCode := -1;
   hmiStns[2].wip[43].pnCode[0] := 0;
   hmiStns[2].wip[43].pnCode[1] := 0;
   hmiStns[2].wip[43].pnCode[2] := 0;
   hmiStns[2].wip[43].pnCode[3] := 0;
   hmiStns[2].wip[43].pnCode[4] := 0;
   hmiStns[2].wip[43].pnCode[5] := 0;
   hmiStns[2].wip[43].pnCode[6] := 0;
   hmiStns[2].wip[43].pnCode[7] := 0;
   hmiStns[2].wip[44].wipCode := -1;
   hmiStns[2].wip[44].pnCode[0] := 0;
   hmiStns[2].wip[44].pnCode[1] := 0;
   hmiStns[2].wip[44].pnCode[2] := 0;
   hmiStns[2].wip[44].pnCode[3] := 0;
   hmiStns[2].wip[44].pnCode[4] := 0;
   hmiStns[2].wip[44].pnCode[5] := 0;
   hmiStns[2].wip[44].pnCode[6] := 0;
   hmiStns[2].wip[44].pnCode[7] := 0;
   hmiStns[2].wip[45].wipCode := -1;
   hmiStns[2].wip[45].pnCode[0] := 0;
   hmiStns[2].wip[45].pnCode[1] := 0;
   hmiStns[2].wip[45].pnCode[2] := 0;
   hmiStns[2].wip[45].pnCode[3] := 0;
   hmiStns[2].wip[45].pnCode[4] := 0;
   hmiStns[2].wip[45].pnCode[5] := 0;
   hmiStns[2].wip[45].pnCode[6] := 0;
   hmiStns[2].wip[45].pnCode[7] := 0;
   hmiStns[2].wip[46].wipCode := -1;
   hmiStns[2].wip[46].pnCode[0] := 0;
   hmiStns[2].wip[46].pnCode[1] := 0;
   hmiStns[2].wip[46].pnCode[2] := 0;
   hmiStns[2].wip[46].pnCode[3] := 0;
   hmiStns[2].wip[46].pnCode[4] := 0;
   hmiStns[2].wip[46].pnCode[5] := 0;
   hmiStns[2].wip[46].pnCode[6] := 0;
   hmiStns[2].wip[46].pnCode[7] := 0;
   hmiStns[2].wip[47].wipCode := -1;
   hmiStns[2].wip[47].pnCode[0] := 0;
   hmiStns[2].wip[47].pnCode[1] := 0;
   hmiStns[2].wip[47].pnCode[2] := 0;
   hmiStns[2].wip[47].pnCode[3] := 0;
   hmiStns[2].wip[47].pnCode[4] := 0;
   hmiStns[2].wip[47].pnCode[5] := 0;
   hmiStns[2].wip[47].pnCode[6] := 0;
   hmiStns[2].wip[47].pnCode[7] := 0;
   hmiStns[2].wip[48].wipCode := -1;
   hmiStns[2].wip[48].pnCode[0] := 0;
   hmiStns[2].wip[48].pnCode[1] := 0;
   hmiStns[2].wip[48].pnCode[2] := 0;
   hmiStns[2].wip[48].pnCode[3] := 0;
   hmiStns[2].wip[48].pnCode[4] := 0;
   hmiStns[2].wip[48].pnCode[5] := 0;
   hmiStns[2].wip[48].pnCode[6] := 0;
   hmiStns[2].wip[48].pnCode[7] := 0;
   hmiStns[2].wip[49].wipCode := -1;
   hmiStns[2].wip[49].pnCode[0] := 0;
   hmiStns[2].wip[49].pnCode[1] := 0;
   hmiStns[2].wip[49].pnCode[2] := 0;
   hmiStns[2].wip[49].pnCode[3] := 0;
   hmiStns[2].wip[49].pnCode[4] := 0;
   hmiStns[2].wip[49].pnCode[5] := 0;
   hmiStns[2].wip[49].pnCode[6] := 0;
   hmiStns[2].wip[49].pnCode[7] := 0;
   hmiStns[3].wip[0].wipCode := 17009;
   hmiStns[3].wip[0].pnCode[0] := 0;
   hmiStns[3].wip[0].pnCode[1] := 243000;
   hmiStns[3].wip[0].pnCode[2] := 52000;
   hmiStns[3].wip[0].pnCode[3] := 0;
   hmiStns[3].wip[0].pnCode[4] := 0;
   hmiStns[3].wip[0].pnCode[5] := 0;
   hmiStns[3].wip[0].pnCode[6] := 31000;
   hmiStns[3].wip[0].pnCode[7] := 73000;
   hmiStns[3].wip[1].wipCode := 69063;
   hmiStns[3].wip[1].pnCode[0] := 0;
   hmiStns[3].wip[1].pnCode[1] := 243000;
   hmiStns[3].wip[1].pnCode[2] := 217000;
   hmiStns[3].wip[1].pnCode[3] := 0;
   hmiStns[3].wip[1].pnCode[4] := 0;
   hmiStns[3].wip[1].pnCode[5] := 0;
   hmiStns[3].wip[1].pnCode[6] := 218000;
   hmiStns[3].wip[1].pnCode[7] := 223000;
   hmiStns[3].wip[2].wipCode := 65047;
   hmiStns[3].wip[2].pnCode[0] := 0;
   hmiStns[3].wip[2].pnCode[1] := 243000;
   hmiStns[3].wip[2].pnCode[2] := 228000;
   hmiStns[3].wip[2].pnCode[3] := 231000;
   hmiStns[3].wip[2].pnCode[4] := 0;
   hmiStns[3].wip[2].pnCode[5] := 229000;
   hmiStns[3].wip[2].pnCode[6] := 227000;
   hmiStns[3].wip[2].pnCode[7] := 230000;
   hmiStns[3].wip[3].wipCode := 68046;
   hmiStns[3].wip[3].pnCode[0] := 0;
   hmiStns[3].wip[3].pnCode[1] := 243000;
   hmiStns[3].wip[3].pnCode[2] := 164000;
   hmiStns[3].wip[3].pnCode[3] := 0;
   hmiStns[3].wip[3].pnCode[4] := 0;
   hmiStns[3].wip[3].pnCode[5] := 165000;
   hmiStns[3].wip[3].pnCode[6] := 202000;
   hmiStns[3].wip[3].pnCode[7] := 203000;
   hmiStns[3].wip[4].wipCode := 64006;
   hmiStns[3].wip[4].pnCode[0] := 0;
   hmiStns[3].wip[4].pnCode[1] := 243000;
   hmiStns[3].wip[4].pnCode[2] := 200000;
   hmiStns[3].wip[4].pnCode[3] := 0;
   hmiStns[3].wip[4].pnCode[4] := 0;
   hmiStns[3].wip[4].pnCode[5] := 201000;
   hmiStns[3].wip[4].pnCode[6] := 202000;
   hmiStns[3].wip[4].pnCode[7] := 203000;
   hmiStns[3].wip[5].wipCode := 66005;
   hmiStns[3].wip[5].pnCode[0] := 0;
   hmiStns[3].wip[5].pnCode[1] := 243000;
   hmiStns[3].wip[5].pnCode[2] := 164000;
   hmiStns[3].wip[5].pnCode[3] := 0;
   hmiStns[3].wip[5].pnCode[4] := 0;
   hmiStns[3].wip[5].pnCode[5] := 165000;
   hmiStns[3].wip[5].pnCode[6] := 202000;
   hmiStns[3].wip[5].pnCode[7] := 203000;
   hmiStns[3].wip[6].wipCode := 67000;
   hmiStns[3].wip[6].pnCode[0] := 0;
   hmiStns[3].wip[6].pnCode[1] := 243000;
   hmiStns[3].wip[6].pnCode[2] := 0;